// TIA Portal project "DnomaidDBMS" (V13) (continued)

   IF #RESET THEN
       #FB_FAULT := FALSE;
       IF #TimerHmiScript.Q THEN
           #NEW := FALSE;
       END_IF;
   END_IF;

   #FB_RET_VAL:=0;
   #NewLog:=FALSE;
   #NewData:="#COMP_DATETIME"(DT1:=#LAST_LOG.DatabaseTable.DateTime , DT2:=#DATE_LAST_LOG); //#COMP_DATETIME GT_DT

   IF #NewData THEN
       FOR #NArray01:=#LOG_LIST_MAX TO #LOG_LIST_MIN BY -1 DO
           IF(#NArray01=#LOG_LIST_MIN AND #LOG_LIST[#NArray01].Request=0)THEN //First position empty
               #NewLog:= TRUE;        
           ELSIF(#NArray01<>#LOG_LIST_MIN AND #LOG_LIST[#NArray01].Request=0)THEN //Next
               IF(#LOG_LIST[#NArray01-1].Request=0)THEN
                   CONTINUE;
               END_IF;    
               #NewLog:=TRUE;                                          
           END_IF;       
           IF(#NewLog)THEN
               #nSec:=1;
               L_00: ;
                   CASE #nSec OF
                   1://---->Copy the log                    
                       #RetVal01:=FILL(BVAL:=#LAST_LOG, BLK=>#LOG_LIST[#NArray01]);
                       GOTO L_IN;
                   2://---->The last date is saved           
                       #RetVal01:=FILL(BVAL:=#LOG_LIST[#NArray01].DatabaseTable.DateTime, BLK=>#DATE_LAST_LOG); 
                       GOTO L_IN;
                   3://---->Pushes the data one position            
                       IF(#NArray01=#LOG_LIST_MAX)THEN
                           #RetVal01:=FILL(BVAL:=#pSourceDB, BLK=>#pDestinationDB);                
                       END_IF; 
                       GOTO L_IN;
                   4://---->Delete last position            
                       IF(#NArray01=#LOG_LIST_MAX)THEN
                           #RetVal01:=FILL(BVAL:=#INI_LOG, BLK=>#LOG_LIST[#LOG_LIST_MAX]);                
                       END_IF; 
                       GOTO L_IN;                                                       
                   ELSE://---->End    
                       GOTO L_EN;
                   END_CASE;
               L_IN://Next
                   IF(#RetVal01<>0)THEN #FB_FAULT:=TRUE; #FB_RET_VAL:=#nSec; GOTO L_EN; END_IF; 
                   #nSec:=#nSec+1; 
                   GOTO L_00;
               L_EN: ;
               EXIT;
           END_IF;                          
       END_FOR;
   END_IF;
   IF #NewData THEN
       #NEW := TRUE;
   END_IF;
END_FUNCTION_BLOCK

FUNCTION_BLOCK "#CTRL_INSERT_DATA"   // FB40, SCL
TITLE = Ctrl insert data
{ S7_Optimized_Access := 'FALSE' }
AUTHOR : QLR
FAMILY : dnomaiD
VERSION : 9.0
BEGIN
   // Timers
   #TimerIni1(IN := #A_TimerIni[1],
               PT := t#1s);
   #Q_TimerIni[1] := #TimerIni1.Q;
   #TimerOutCase1(IN := #A_TimerOutCase[1],
              PT := t#35s);
   #Q_TimerOutCase[1] := #TimerOutCase1.Q;

   #TimerIni2(IN := #A_TimerIni[2],
              PT := t#1s);
   #Q_TimerIni[2] := #TimerIni2.Q;
   #TimerOutCase2(IN := #A_TimerOutCase[2],
                  PT := t#35s);
   #Q_TimerOutCase[2] := #TimerOutCase2.Q;
   #TimerIni := FALSE;
   FOR #"Counter" := #ArrayIni TO #ArrayEnd DO
       IF #A_TimerIni[#"Counter"] THEN
           #TimerIni := TRUE;
       END_IF;
   END_FOR;

   FOR #"Counter" := #ArrayIni TO #ArrayEnd DO

       IF #Q_TimerOutCase[#"Counter"] THEN
           #Status[#"Counter"] := 99;
       END_IF;

       CASE #Status[#"Counter"] OF
           1:  //Ini..
               IF NOT #InsertBarcode[#"Counter"] AND NOT #ResponseInsertCompleted AND #Q_TimerIni[#"Counter"] AND NOT #Reset THEN
                   #Status[#"Counter"] := 1 + #Status[#"Counter"];
               END_IF;
               GOTO END;
           2:  //Waiting for permission to insert data
               IF #InsertPerm THEN
                   #Status[#"Counter"] := 1 + #Status[#"Counter"];
               END_IF;
               GOTO END;
           3:  //Ready
               IF #InsertBarcode[#"Counter"]  THEN
                  #Status[#"Counter"] := 1 + #Status[#"Counter"];
               END_IF;
               GOTO END;
           4:  //Start
               IF NOT #ResponseInsertCompleted AND NOT #InProgress THEN
                   UMOVE_BLK(IN := #DataBarcodeCode[#"Counter"].Digit[1],
                             COUNT := 13,
                             OUT => #DataCode.Digit[1]);
                   #DataScanner.Number := #DataBarcodeScanner[#"Counter"].Number;
                   #InProgress := TRUE;
                   #Status[#"Counter"] := 1 + #Status[#"Counter"];
               END_IF;
               GOTO END;
           5:  // data copied!  
               IF NOT #ResponseInsertCompleted THEN
                   #Insert := TRUE;
                   #Status[#"Counter"] := 1 + #Status[#"Counter"];
               END_IF;
               GOTO END;
           6:  //in progress...
               IF #ResponseInsertCompleted THEN
                   #Insert := FALSE;
                   #InProgress := FALSE;
                   #Status[#"Counter"] := 0;
               END_IF;
               GOTO END;
           99: // time out
               IF #Reset THEN
                   #Insert := FALSE;
                   #InProgress := FALSE;
                   #Status[#"Counter"] := 0;
               END_IF;
           ELSE  
               #Status[#"Counter"] := 1;
               #Insert := FALSE;
               GOTO END;
       END_CASE;
       END: ;

       IF #Status[#"Counter"] = 1 THEN
           IF NOT #InProgress AND NOT #TimerIni THEN
               #A_TimerIni[#"Counter"] := TRUE;
           END_IF;
       ELSE
           #A_TimerIni[#"Counter"] := FALSE;
       END_IF;
       IF #InProgress THEN
           #A_TimerOutCase[#"Counter"] := TRUE;
       ELSE
           #A_TimerOutCase[#"Counter"] := FALSE;
       END_IF;

   END_FOR;
END_FUNCTION_BLOCK

FUNCTION_BLOCK "#SIMU_BARCODE EAN-13"   // FB401, STL
TITLE = Simu Barcode
{ S7_Optimized_Access := 'FALSE' }
AUTHOR : QLR
FAMILY : dnomaiD
VERSION : 9.0
BEGIN

REGION Network 1: Start
         TAR1  #SaveAR1;
         L     STW;
         T     #SaveSTW;
         CLR;
         =     #ValNeg;
         =     #RequestInsert;
         L     0;
         T     #QuaChar;
         T     #BcdSDL4;
         T     #NumDB;

         L     #CodeNum;
         L     #MaxNumber;
         >=I;
         JC    aA01;
         JU    aAFF;
   aA01: NOP   0;
         L     0;
         T     #CodeNum;
         JU    aAFF;
   aAFF: NOP   0;
END_REGION

REGION Network 2: Next
         A     #NextNumber;
         FP    #FpNext;
         JC    cA01;
         JU    END;
   cA01: NOP   0;
         CALL  FILL_BLK
         ( IN    := '0',
           COUNT := #LengthChar,
           OUT   := #CODE.Digit[1]
         );
         L     #CodeNum;
         +     1;
         T     #CodeNum;
         SET;
         S     #RequestInsert;
END_REGION

REGION Network 3: Convert int to char
         L     #""Address_25";
         LAR1;
         L     W[AR1, P#0.0];
         T     #NumDB;
         OPN   DB[ #NumDB];
         L     D[AR1, P#2.0];
         LAR1;
         L     #CodeNum;
         L     0;
         +I;
         JP    BC01;
         JZ    BC02;
         SET;
         =     #ValNeg;
         L     1;
         T     #CodeNum;
         JU    END;
   BC01: NOP   0;  // <0
         ITD;
         DTR;
         ABS;
         LN;
         L     2.302585;
         /R;
         TRUNC;
   BC02: NOP   0;  // ==0
         +     1;
         T     #QuaChar;
         +     1;
         L     #LengthChar;
         >I;
         JC    END;
         TAK;
         L     #CodeNum;
         ITD;
         DTB;
         T     #BcdSDL4;
         L     #BcdSDL4;
         SLD   4;
         T     #BcdSDL4;
         L     #LengthChar;
         L     -1;
         +I;
         L     8;
         *I;
         +AR1;
         L     #QuaChar;
   BC03: NOP   0;  // Loop
         T     #QuaChar;
         L     #BcdSDL4;
         SRD   4;
         T     #BcdSDL4;
         AD    16#0000_000F;
         L     B#16#30;
         OW;
         T     B [ AR1 , P#0.0 ];
         L     DINT#-8;
         +AR1;
         L     #QuaChar;
         LOOP  BC03;
         L     #ScannerNumber;
         T     #ScannerNumberAuto;
END_REGION

REGION Network 4: End
         JU    END;
   END:  NOP   0;
         LAR1  #SaveAR1;
         L     #SaveSTW;
         T     STW;
         SET;
         SAVE;
         BE;
END_REGION
END_FUNCTION_BLOCK

FUNCTION "DATABASE_MANAGER" : Void   // FC30, LAD
TITLE = Database manager
{ S7_Optimized_Access := 'FALSE' }
AUTHOR : QLR
FAMILY : dnomaiD
VERSION : 9.0
   VAR_TEMP   // added for the SCL form of the ladder/FBD networks
      _w1 : Bool;
      _w2 : Bool;
   END_VAR
BEGIN

REGION Network 1: Ctrl insert data Auto
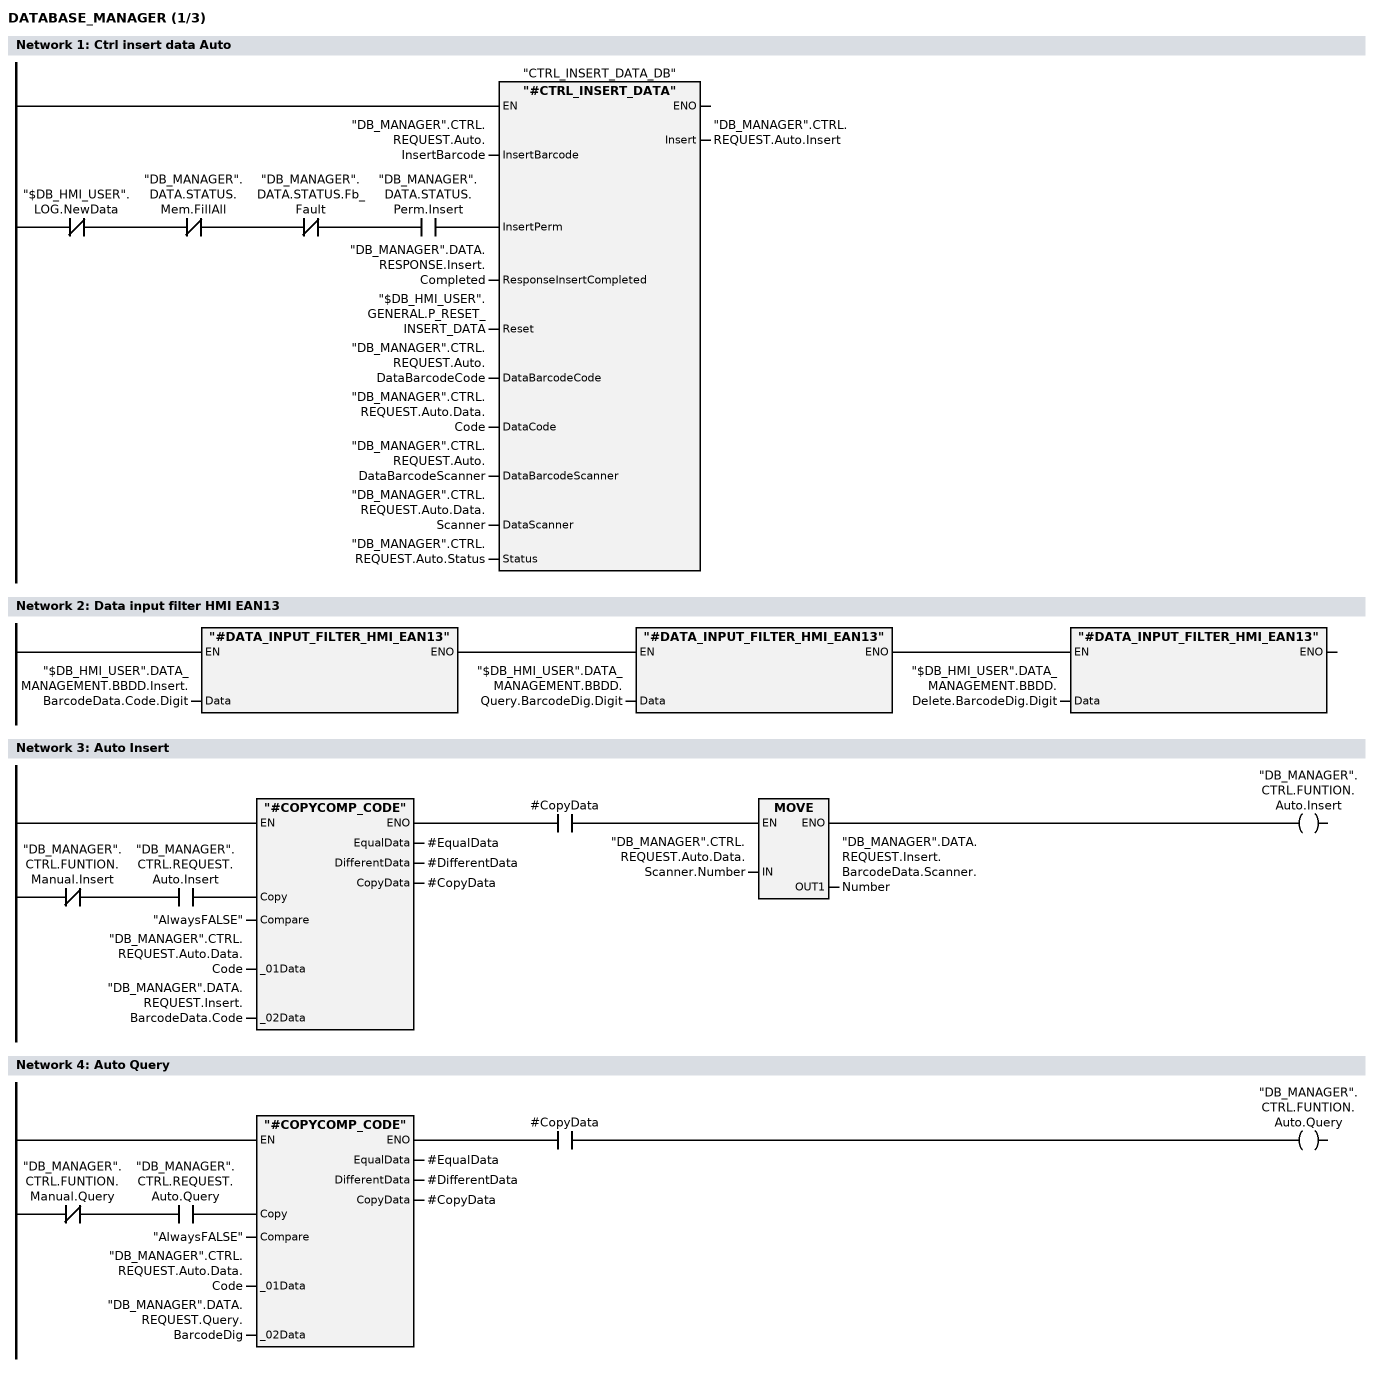
   RUNG wire#powerrail
      "CTRL_INSERT_DATA_DB"(InsertPerm := wire#w1, InsertBarcode := "DB_MANAGER".CTRL.REQUEST.Auto.InsertBarcode, ResponseInsertCompleted := "DB_MANAGER".DATA.RESPONSE.Insert.Completed, Reset := "$DB_HMI_USER".GENERAL.P_RESET_INSERT_DATA, DataBarcodeCode := "DB_MANAGER".CTRL.REQUEST.Auto.DataBarcodeCode, DataCode := "DB_MANAGER".CTRL.REQUEST.Auto.Data.Code, DataBarcodeScanner := "DB_MANAGER".CTRL.REQUEST.Auto.DataBarcodeScanner, DataScanner := "DB_MANAGER".CTRL.REQUEST.Auto.Data.Scanner, Status := "DB_MANAGER".CTRL.REQUEST.Auto.Status, Insert => "DB_MANAGER".CTRL.REQUEST.Auto.Insert)
   END_RUNG
   RUNG wire#powerrail
      I_Contact( "$DB_HMI_USER".LOG.NewData )
      I_Contact( "DB_MANAGER".DATA.STATUS.Mem.FillAll )
      I_Contact( "DB_MANAGER".DATA.STATUS.Fb_Fault )
      Contact( "DB_MANAGER".DATA.STATUS.Perm.Insert )
   END_RUNG wire#w1
   // the same network as SCL:
   "CTRL_INSERT_DATA_DB"(InsertBarcode := "DB_MANAGER".CTRL.REQUEST.Auto.InsertBarcode,   // "#CTRL_INSERT_DATA"
                         InsertPerm := NOT "$DB_HMI_USER".LOG.NewData AND NOT "DB_MANAGER".DATA.STATUS.Mem.FillAll AND NOT "DB_MANAGER".DATA.STATUS.Fb_Fault AND "DB_MANAGER".DATA.STATUS.Perm.Insert,
                         ResponseInsertCompleted := "DB_MANAGER".DATA.RESPONSE.Insert.Completed,
                         Reset := "$DB_HMI_USER".GENERAL.P_RESET_INSERT_DATA,
                         DataBarcodeCode := "DB_MANAGER".CTRL.REQUEST.Auto.DataBarcodeCode,
                         DataCode := "DB_MANAGER".CTRL.REQUEST.Auto.Data.Code,
                         DataBarcodeScanner := "DB_MANAGER".CTRL.REQUEST.Auto.DataBarcodeScanner,
                         DataScanner := "DB_MANAGER".CTRL.REQUEST.Auto.Data.Scanner,
                         Status := "DB_MANAGER".CTRL.REQUEST.Auto.Status,
                         Insert => "DB_MANAGER".CTRL.REQUEST.Auto.Insert);
END_REGION

REGION Network 2: Data input filter HMI EAN13
   RUNG wire#powerrail
      "#DATA_INPUT_FILTER_HMI_EAN13"(Data := "$DB_HMI_USER".DATA_MANAGEMENT.BBDD.Insert.BarcodeData.Code.Digit)
      "#DATA_INPUT_FILTER_HMI_EAN13"(Data := "$DB_HMI_USER".DATA_MANAGEMENT.BBDD.Query.BarcodeDig.Digit)
      "#DATA_INPUT_FILTER_HMI_EAN13"(Data := "$DB_HMI_USER".DATA_MANAGEMENT.BBDD.Delete.BarcodeDig.Digit)
   END_RUNG
   // the same network as SCL:
   "#DATA_INPUT_FILTER_HMI_EAN13"(Data := "$DB_HMI_USER".DATA_MANAGEMENT.BBDD.Insert.BarcodeData.Code.Digit,
                           ENO => #_w1);
   "#DATA_INPUT_FILTER_HMI_EAN13"(EN := #_w1,
                           Data := "$DB_HMI_USER".DATA_MANAGEMENT.BBDD.Query.BarcodeDig.Digit,
                           ENO => #_w2);
   IF #_w2 THEN
       "#DATA_INPUT_FILTER_HMI_EAN13"(Data := "$DB_HMI_USER".DATA_MANAGEMENT.BBDD.Delete.BarcodeDig.Digit);
   END_IF;
END_REGION

REGION Network 3: Auto Insert
   RUNG wire#powerrail
      "#COPYCOMP_CODE"(Copy := wire#w1, Compare := "AlwaysFALSE", _01Data := "DB_MANAGER".CTRL.REQUEST.Auto.Data.Code, _02Data := "DB_MANAGER".DATA.REQUEST.Insert.BarcodeData.Code, EqualData => #EqualData, DifferentData => #DifferentData, CopyData => #CopyData)
      Contact( #CopyData )
      { S7_GenerateENO := "TRUE" } Move(in := "DB_MANAGER".CTRL.REQUEST.Auto.Data.Scanner.Number, out1 => "DB_MANAGER".DATA.REQUEST.Insert.BarcodeData.Scanner.Number)
      Coil( "DB_MANAGER".CTRL.FUNTION.Auto.Insert )
   END_RUNG
   RUNG wire#powerrail
      I_Contact( "DB_MANAGER".CTRL.FUNTION.Manual.Insert )
      Contact( "DB_MANAGER".CTRL.REQUEST.Auto.Insert )
   END_RUNG wire#w1
   // the same network as SCL:
   // ENO of a box is taken as its EN; it also drops when the box reports an error
   "#COPYCOMP_CODE"(Copy := NOT "DB_MANAGER".CTRL.FUNTION.Manual.Insert AND "DB_MANAGER".CTRL.REQUEST.Auto.Insert,
                    Compare := "AlwaysFALSE",
                    _01Data := "DB_MANAGER".CTRL.REQUEST.Auto.Data.Code,
                    _02Data := "DB_MANAGER".DATA.REQUEST.Insert.BarcodeData.Code,
                    EqualData => #EqualData,
                    DifferentData => #DifferentData,
                    CopyData => #CopyData,
                    ENO => #_w1);
   #_w2 := #_w1 AND #CopyData;
   IF #_w2 THEN
       "DB_MANAGER".DATA.REQUEST.Insert.BarcodeData.Scanner.Number := "DB_MANAGER".CTRL.REQUEST.Auto.Data.Scanner.Number;
   END_IF;
   "DB_MANAGER".CTRL.FUNTION.Auto.Insert := #_w2;
END_REGION

REGION Network 4: Auto Query
   RUNG wire#powerrail
      "#COPYCOMP_CODE"(Copy := wire#w1, Compare := "AlwaysFALSE", _01Data := "DB_MANAGER".CTRL.REQUEST.Auto.Data.Code, _02Data := "DB_MANAGER".DATA.REQUEST.Query.BarcodeDig, EqualData => #EqualData, DifferentData => #DifferentData, CopyData => #CopyData)
      Contact( #CopyData )
      Coil( "DB_MANAGER".CTRL.FUNTION.Auto.Query )
   END_RUNG
   RUNG wire#powerrail
      I_Contact( "DB_MANAGER".CTRL.FUNTION.Manual.Query )
      Contact( "DB_MANAGER".CTRL.REQUEST.Auto.Query )
   END_RUNG wire#w1
   // the same network as SCL:
   "#COPYCOMP_CODE"(Copy := NOT "DB_MANAGER".CTRL.FUNTION.Manual.Query AND "DB_MANAGER".CTRL.REQUEST.Auto.Query,
                    Compare := "AlwaysFALSE",
                    _01Data := "DB_MANAGER".CTRL.REQUEST.Auto.Data.Code,
                    _02Data := "DB_MANAGER".DATA.REQUEST.Query.BarcodeDig,
                    EqualData => #EqualData,
                    DifferentData => #DifferentData,
                    CopyData => #CopyData,
                    ENO => #_w1);
   "DB_MANAGER".CTRL.FUNTION.Auto.Query := #_w1 AND #CopyData;
END_REGION

REGION Network 5: Auto Delete
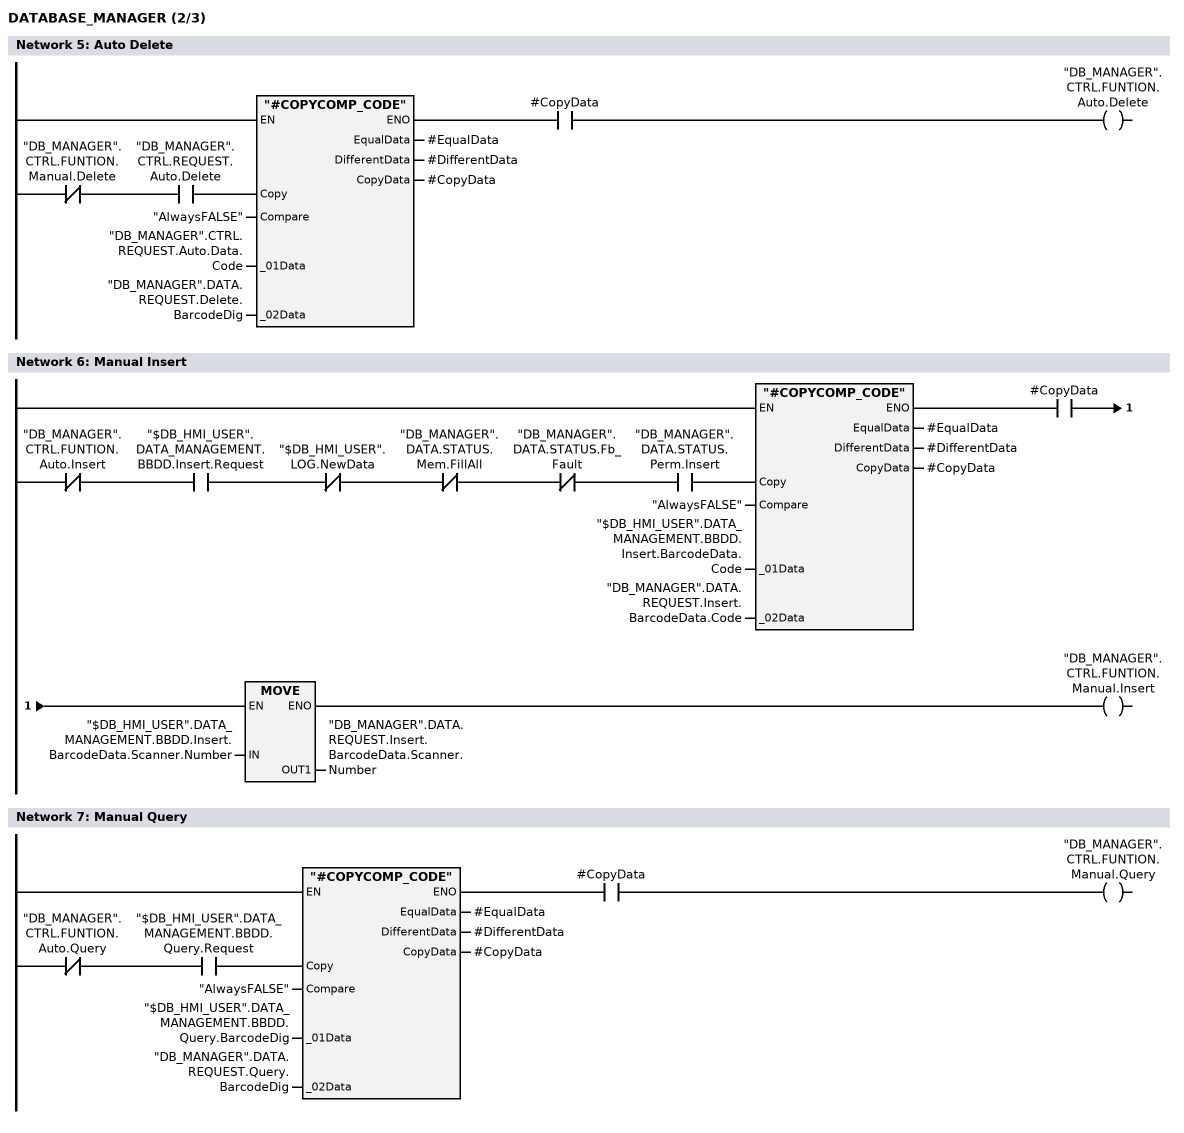
   RUNG wire#powerrail
      "#COPYCOMP_CODE"(Copy := wire#w1, Compare := "AlwaysFALSE", _01Data := "DB_MANAGER".CTRL.REQUEST.Auto.Data.Code, _02Data := "DB_MANAGER".DATA.REQUEST.Delete.BarcodeDig, EqualData => #EqualData, DifferentData => #DifferentData, CopyData => #CopyData)
      Contact( #CopyData )
      Coil( "DB_MANAGER".CTRL.FUNTION.Auto.Delete )
   END_RUNG
   RUNG wire#powerrail
      I_Contact( "DB_MANAGER".CTRL.FUNTION.Manual.Delete )
      Contact( "DB_MANAGER".CTRL.REQUEST.Auto.Delete )
   END_RUNG wire#w1
   // the same network as SCL:
   "#COPYCOMP_CODE"(Copy := NOT "DB_MANAGER".CTRL.FUNTION.Manual.Delete AND "DB_MANAGER".CTRL.REQUEST.Auto.Delete,
                    Compare := "AlwaysFALSE",
                    _01Data := "DB_MANAGER".CTRL.REQUEST.Auto.Data.Code,
                    _02Data := "DB_MANAGER".DATA.REQUEST.Delete.BarcodeDig,
                    EqualData => #EqualData,
                    DifferentData => #DifferentData,
                    CopyData => #CopyData,
                    ENO => #_w1);
   "DB_MANAGER".CTRL.FUNTION.Auto.Delete := #_w1 AND #CopyData;
END_REGION

REGION Network 6: Manual Insert
   RUNG wire#powerrail
      "#COPYCOMP_CODE"(Copy := wire#w1, Compare := "AlwaysFALSE", _01Data := "$DB_HMI_USER".DATA_MANAGEMENT.BBDD.Insert.BarcodeData.Code, _02Data := "DB_MANAGER".DATA.REQUEST.Insert.BarcodeData.Code, EqualData => #EqualData, DifferentData => #DifferentData, CopyData => #CopyData)
      Contact( #CopyData )
      { S7_GenerateENO := "TRUE" } Move(in := "$DB_HMI_USER".DATA_MANAGEMENT.BBDD.Insert.BarcodeData.Scanner.Number, out1 => "DB_MANAGER".DATA.REQUEST.Insert.BarcodeData.Scanner.Number)
      Coil( "DB_MANAGER".CTRL.FUNTION.Manual.Insert )
   END_RUNG
   RUNG wire#powerrail
      I_Contact( "DB_MANAGER".CTRL.FUNTION.Auto.Insert )
      Contact( "$DB_HMI_USER".DATA_MANAGEMENT.BBDD.Insert.Request )
      I_Contact( "$DB_HMI_USER".LOG.NewData )
      I_Contact( "DB_MANAGER".DATA.STATUS.Mem.FillAll )
      I_Contact( "DB_MANAGER".DATA.STATUS.Fb_Fault )
      Contact( "DB_MANAGER".DATA.STATUS.Perm.Insert )
   END_RUNG wire#w1
   // the same network as SCL:
   // ENO of a box is taken as its EN; it also drops when the box reports an error
   "#COPYCOMP_CODE"(Copy := NOT "DB_MANAGER".CTRL.FUNTION.Auto.Insert AND "$DB_HMI_USER".DATA_MANAGEMENT.BBDD.Insert.Request AND NOT "$DB_HMI_USER".LOG.NewData AND NOT "DB_MANAGER".DATA.STATUS.Mem.FillAll AND NOT "DB_MANAGER".DATA.STATUS.Fb_Fault AND "DB_MANAGER".DATA.STATUS.Perm.Insert,
                    Compare := "AlwaysFALSE",
                    _01Data := "$DB_HMI_USER".DATA_MANAGEMENT.BBDD.Insert.BarcodeData.Code,
                    _02Data := "DB_MANAGER".DATA.REQUEST.Insert.BarcodeData.Code,
                    EqualData => #EqualData,
                    DifferentData => #DifferentData,
                    CopyData => #CopyData,
                    ENO => #_w1);
   #_w2 := #_w1 AND #CopyData;
   IF #_w2 THEN
       "DB_MANAGER".DATA.REQUEST.Insert.BarcodeData.Scanner.Number := "$DB_HMI_USER".DATA_MANAGEMENT.BBDD.Insert.BarcodeData.Scanner.Number;
   END_IF;
   "DB_MANAGER".CTRL.FUNTION.Manual.Insert := #_w2;
END_REGION

REGION Network 7: Manual Query
   RUNG wire#powerrail
      "#COPYCOMP_CODE"(Copy := wire#w1, Compare := "AlwaysFALSE", _01Data := "$DB_HMI_USER".DATA_MANAGEMENT.BBDD.Query.BarcodeDig, _02Data := "DB_MANAGER".DATA.REQUEST.Query.BarcodeDig, EqualData => #EqualData, DifferentData => #DifferentData, CopyData => #CopyData)
      Contact( #CopyData )
      Coil( "DB_MANAGER".CTRL.FUNTION.Manual.Query )
   END_RUNG
   RUNG wire#powerrail
      I_Contact( "DB_MANAGER".CTRL.FUNTION.Auto.Query )
      Contact( "$DB_HMI_USER".DATA_MANAGEMENT.BBDD.Query.Request )
   END_RUNG wire#w1
   // the same network as SCL:
   "#COPYCOMP_CODE"(Copy := NOT "DB_MANAGER".CTRL.FUNTION.Auto.Query AND "$DB_HMI_USER".DATA_MANAGEMENT.BBDD.Query.Request,
                    Compare := "AlwaysFALSE",
                    _01Data := "$DB_HMI_USER".DATA_MANAGEMENT.BBDD.Query.BarcodeDig,
                    _02Data := "DB_MANAGER".DATA.REQUEST.Query.BarcodeDig,
                    EqualData => #EqualData,
                    DifferentData => #DifferentData,
                    CopyData => #CopyData,
                    ENO => #_w1);
   "DB_MANAGER".CTRL.FUNTION.Manual.Query := #_w1 AND #CopyData;
END_REGION

REGION Network 8: Manual Delete
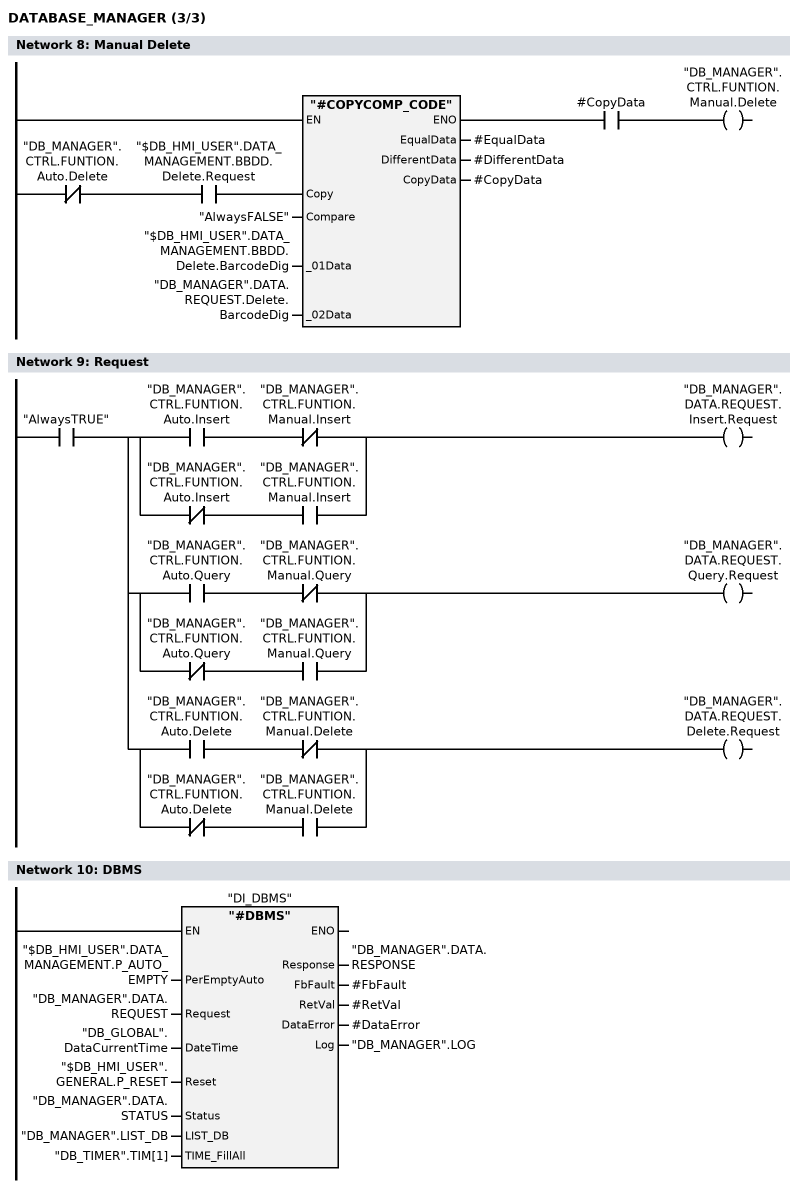
   RUNG wire#powerrail
      "#COPYCOMP_CODE"(Copy := wire#w1, Compare := "AlwaysFALSE", _01Data := "$DB_HMI_USER".DATA_MANAGEMENT.BBDD.Delete.BarcodeDig, _02Data := "DB_MANAGER".DATA.REQUEST.Delete.BarcodeDig, EqualData => #EqualData, DifferentData => #DifferentData, CopyData => #CopyData)
      Contact( #CopyData )
      Coil( "DB_MANAGER".CTRL.FUNTION.Manual.Delete )
   END_RUNG
   RUNG wire#powerrail
      I_Contact( "DB_MANAGER".CTRL.FUNTION.Auto.Delete )
      Contact( "$DB_HMI_USER".DATA_MANAGEMENT.BBDD.Delete.Request )
   END_RUNG wire#w1
   // the same network as SCL:
   "#COPYCOMP_CODE"(Copy := NOT "DB_MANAGER".CTRL.FUNTION.Auto.Delete AND "$DB_HMI_USER".DATA_MANAGEMENT.BBDD.Delete.Request,
                    Compare := "AlwaysFALSE",
                    _01Data := "$DB_HMI_USER".DATA_MANAGEMENT.BBDD.Delete.BarcodeDig,
                    _02Data := "DB_MANAGER".DATA.REQUEST.Delete.BarcodeDig,
                    EqualData => #EqualData,
                    DifferentData => #DifferentData,
                    CopyData => #CopyData,
                    ENO => #_w1);
   "DB_MANAGER".CTRL.FUNTION.Manual.Delete := #_w1 AND #CopyData;
END_REGION

REGION Network 9: Request
   RUNG wire#powerrail
      Contact( "AlwaysTRUE" )
      wire#w1
      Contact( "DB_MANAGER".CTRL.FUNTION.Auto.Insert )
      I_Contact( "DB_MANAGER".CTRL.FUNTION.Manual.Insert )
      wire#w2
      Coil( "DB_MANAGER".DATA.REQUEST.Insert.Request )
   END_RUNG
   RUNG wire#w1
      I_Contact( "DB_MANAGER".CTRL.FUNTION.Auto.Insert )
      Contact( "DB_MANAGER".CTRL.FUNTION.Manual.Insert )
   END_RUNG wire#w2
   RUNG wire#w1
      Contact( "DB_MANAGER".CTRL.FUNTION.Auto.Query )
      I_Contact( "DB_MANAGER".CTRL.FUNTION.Manual.Query )
      wire#w3
      Coil( "DB_MANAGER".DATA.REQUEST.Query.Request )
   END_RUNG
   RUNG wire#w1
      I_Contact( "DB_MANAGER".CTRL.FUNTION.Auto.Query )
      Contact( "DB_MANAGER".CTRL.FUNTION.Manual.Query )
   END_RUNG wire#w3
   RUNG wire#w1
      Contact( "DB_MANAGER".CTRL.FUNTION.Auto.Delete )
      I_Contact( "DB_MANAGER".CTRL.FUNTION.Manual.Delete )
      wire#w4
      Coil( "DB_MANAGER".DATA.REQUEST.Delete.Request )
   END_RUNG
   RUNG wire#w1
      I_Contact( "DB_MANAGER".CTRL.FUNTION.Auto.Delete )
      Contact( "DB_MANAGER".CTRL.FUNTION.Manual.Delete )
   END_RUNG wire#w4
   // the same network as SCL:
   "DB_MANAGER".DATA.REQUEST.Insert.Request := "AlwaysTRUE" AND (("DB_MANAGER".CTRL.FUNTION.Auto.Insert AND NOT "DB_MANAGER".CTRL.FUNTION.Manual.Insert) OR (NOT "DB_MANAGER".CTRL.FUNTION.Auto.Insert AND "DB_MANAGER".CTRL.FUNTION.Manual.Insert));
   "DB_MANAGER".DATA.REQUEST.Query.Request := "AlwaysTRUE" AND (("DB_MANAGER".CTRL.FUNTION.Auto.Query AND NOT "DB_MANAGER".CTRL.FUNTION.Manual.Query) OR (NOT "DB_MANAGER".CTRL.FUNTION.Auto.Query AND "DB_MANAGER".CTRL.FUNTION.Manual.Query));
   "DB_MANAGER".DATA.REQUEST.Delete.Request := "AlwaysTRUE" AND (("DB_MANAGER".CTRL.FUNTION.Auto.Delete AND NOT "DB_MANAGER".CTRL.FUNTION.Manual.Delete) OR (NOT "DB_MANAGER".CTRL.FUNTION.Auto.Delete AND "DB_MANAGER".CTRL.FUNTION.Manual.Delete));
END_REGION

REGION Network 10: DBMS
   RUNG wire#powerrail
      "DI_DBMS"(PerEmptyAuto := "$DB_HMI_USER".DATA_MANAGEMENT.P_AUTO_EMPTY, Request := "DB_MANAGER".DATA.REQUEST, DateTime := "DB_GLOBAL".DataCurrentTime, Reset := "$DB_HMI_USER".GENERAL.P_RESET, Status := "DB_MANAGER".DATA.STATUS, LIST_DB := "DB_MANAGER".LIST_DB, TIME_FillAll := "DB_TIMER".TIM[1], Response => "DB_MANAGER".DATA.RESPONSE, FbFault => #FbFault, RetVal => #RetVal, DataError => #DataError, Log => "DB_MANAGER".LOG)
   END_RUNG
   // the same network as SCL:
   "DI_DBMS"(PerEmptyAuto := "$DB_HMI_USER".DATA_MANAGEMENT.P_AUTO_EMPTY,   // "#DBMS"
             Request := "DB_MANAGER".DATA.REQUEST,
             DateTime := "DB_GLOBAL".DataCurrentTime,
             Reset := "$DB_HMI_USER".GENERAL.P_RESET,
             Status := "DB_MANAGER".DATA.STATUS,
             LIST_DB := "DB_MANAGER".LIST_DB,
             TIME_FillAll := "DB_TIMER".TIM[1],
             Response => "DB_MANAGER".DATA.RESPONSE,
             FbFault => #FbFault,
             RetVal => #RetVal,
             DataError => #DataError,
             Log => "DB_MANAGER".LOG);
END_REGION

REGION Network 11 (STL): End
         SET;
         SAVE;
         BE;
END_REGION
END_FUNCTION

FUNCTION "#COPYCOMP_CODE" : Void   // FC302, STL
TITLE = Copy||Compare
{ S7_Optimized_Access := 'FALSE' }
AUTHOR : QLR
FAMILY : dnomaiD
VERSION : 9.0
BEGIN

REGION Network 1: Home
         TAR1  #SaveAR1;
         TAR2  #SaveAR2;
         L     STW;
         T     #SaveSTW;

         SET;
         R     #EqualData;
         R     #DifferentData;
         R     #CopyData;

         L     #""Address_11";
         L     #""Address_3";
         XOD;
         L     8;
         /D;
         T     #Long;
         L     P#1.0;
         T     #LongAR;

         L     #""Address_44";
         LAR1;
         L     LW [ AR1 , P#0.0 ];
         T     #NumDB01;
         L     LW [ AR1 , P#4.0 ];
         LAR1;
         OPN   DB [ #NumDB01 ];

         L     #""Address_42";
         LAR2;
         L     LW [ AR2 , P#0.0 ];
         T     #NumDB02;
         L     LW [ AR2 , P#4.0 ];
         LAR2;
         OPN   DI [ #NumDB02];
END_REGION

REGION Network 2: Copy
         AN    #Copy;
         JC    COWF;
         L     #Long;
   COW0: NOP   0;
         T     #Counter01;
         L     DBB[AR1, P#0.0];
         T     DIB[AR2, P#0.0];
         L     #LongAR;
         +AR1;
         +AR2;
         L     #Counter01;
         LOOP  COW0;
         SET;
         S     #CopyData;
         S     #EqualData;
         JU    END;
   COWF: NOP   0;
         SET;
         R     #CopyData;
         JU    COFF;
   COFF: NOP   0;
END_REGION

REGION Network 3: Compare
         AN    #Compare;
         JC    CMWF;
         L     #Long;
   CM00: NOP   0;
         T     #Counter01;
         L     DBB[AR1, P#0.0];
         L     DIB[AR2, P#0.0];
         <>I;
         JC    CM01;
         L     #LongAR;
         +AR1;
         +AR2;
         L     #Counter01;
         LOOP  CM00;
         SET;
         S     #EqualData;
         R     #DifferentData;
         JU    CMFF;
         JU    CM01;
   CM01: NOP   0;
         SET;
         R     #EqualData;
         S     #DifferentData;
         JU    CMFF;
         JU    CMWF;
   CMWF: NOP   0;
         SET;
         R     #EqualData;
         R     #DifferentData;
         JU    CMFF;
   CMFF: NOP   0;
END_REGION

REGION Network 4: End
         JU    END;
   END:  NOP   0;
         LAR1  #SaveAR1;
         LAR2  #SaveAR2;
         L     #SaveSTW;
         T     STW;
         SET;
         SAVE;
         BE;
END_REGION
END_FUNCTION

FUNCTION "#COMP_DATETIME" : Void   // FC304, STL
TITLE = Compare DT1>DT2
{ S7_Optimized_Access := 'FALSE' }
AUTHOR : QLR
FAMILY : dnomaiD
VERSION : 9.0
BEGIN

REGION Network 1: Start
         L     STW;
         T     #SaveSTW;
         L     0;
         T     #DB1;
         T     #DB2;
         T     #AuxYearDt;
         T     #YearDt1;
         T     #YearDt2;
         T     #Loop1;
         T     #Loop2;
END_REGION

REGION Network 2: Pointer
         L     #""Address_8";
         LAR1;
         L     #""Address_10";
         LAR2;
         L     W[AR1, P#0.0];
         T     #DB1;
         OPN   DB [ #DB1];
         L     D[AR1, P#2.0];
         LAR1;
         L     W[AR2, P#0.0];
         T     #DB2;
         OPN   DI [ #DB2];
         L     D[AR2, P#2.0];
         OD    16#0100_0000;
         LAR2;
         SET;
         SAVE;
END_REGION

REGION Network 3: Check if it is a BCD number
         JU    DT00;
         L     1;
         T     #Loop1;
   DT00: NOP   0;
         L     #Loop1;
         JL    DTXX;
         JU    DT01;  //Data time 1
         JU    DT02;  //Data time 2
   DTXX: JU    DTFF;  //End
   DT01: NOP   0;
         L     B[AR1, P#0.0];
         T     #YearDt1;
         T     #AuxYearDt;
         JU    DTXF;
   DT02: NOP   0;
         L     B[AR2, P#0.0];
         T     #YearDt2;
         T     #AuxYearDt;
         JU    DTXF;
   DTXF: NOP   0;
         AW    16#6666;
         PUSH;
         JZ    DTOK;
         SLW   1;
         L     #AuxYearDt;
         AW;
         AW    16#8888;
         JN    ERR;
         TAK;
         AW    16#4444;
         SLW   1;
         L     #AuxYearDt;
         AW;
         JN    ERR;
   DTOK: NOP   0;
         L     #Loop1;
         +     1;
         T     #Loop1;
         JU    DT00;
         JU    DTFF;
   DTFF: NOP   0;
END_REGION

REGION Network 4: Year
         JU    YEAR;
   YEAR: NOP   0;
         L     89;
         L     #YearDt1;  //(1990-1999)
         BTI;
         <I;
         JC    YE1;
         +     100;  //(2000-2089)
   YE1:  NOP   0;
         T     #YearDt1;
         L     89;
         L     #YearDt2;  //(1990-1999)
         BTI;
         <I;
         JC    YE2;
         +     100;  //(2000-2089)
   YE2:  NOP   0;
         T     #YearDt2;
         L     #YearDt1;
         <I;
         JC    SET;
         >I;
         JC    RESE;
END_REGION

